   END_RUNG
   RUNG wire#w1
      Contact( %DB67.DBX7.1 )
      R_Coil( %DB60.DBX7.1 )
   END_RUNG
   RUNG wire#w1
      Contact( %DB67.DBX7.2 )
      R_Coil( %DB60.DBX7.2 )
   END_RUNG
   RUNG wire#w1
      Contact( %DB67.DBX7.3 )
      R_Coil( %DB60.DBX7.3 )
   END_RUNG
   RUNG wire#w1
      Contact( %DB67.DBX7.4 )
      R_Coil( %DB60.DBX7.4 )
   END_RUNG
   RUNG wire#w1
      Contact( %DB67.DBX7.5 )
      R_Coil( %DB60.DBX7.5 )
   END_RUNG
   RUNG wire#w1
      Contact( %DB67.DBX7.6 )
      R_Coil( %DB60.DBX7.6 )
   END_RUNG
   RUNG wire#w1
      Contact( %DB67.DBX7.7 )
      R_Coil( %DB60.DBX7.7 )
   END_RUNG
   // the same network as SCL:
   IF "AlwaysFALSE" AND %DB67.DBX0.0 THEN %DB60.DBX0.0 := FALSE; END_IF;
   IF "AlwaysFALSE" AND %DB67.DBX0.1 THEN %DB60.DBX0.1 := FALSE; END_IF;
   IF "AlwaysFALSE" AND %DB67.DBX0.2 THEN %DB60.DBX0.2 := FALSE; END_IF;
   IF "AlwaysFALSE" AND %DB67.DBX0.3 THEN %DB60.DBX0.3 := FALSE; END_IF;
   IF "AlwaysFALSE" AND %DB67.DBX0.4 THEN %DB60.DBX0.4 := FALSE; END_IF;
   IF "AlwaysFALSE" AND %DB67.DBX0.5 THEN %DB60.DBX0.5 := FALSE; END_IF;
   IF "AlwaysFALSE" AND %DB67.DBX0.6 THEN %DB60.DBX0.6 := FALSE; END_IF;
   IF "AlwaysFALSE" AND %DB67.DBX0.7 THEN %DB60.DBX0.7 := FALSE; END_IF;
   IF "AlwaysFALSE" AND %DB67.DBX1.0 THEN %DB60.DBX1.0 := FALSE; END_IF;
   IF "AlwaysFALSE" AND %DB67.DBX1.1 THEN %DB60.DBX1.1 := FALSE; END_IF;
   IF "AlwaysFALSE" AND %DB67.DBX1.2 THEN %DB60.DBX1.2 := FALSE; END_IF;
   IF "AlwaysFALSE" AND %DB67.DBX1.3 THEN %DB60.DBX1.3 := FALSE; END_IF;
   IF "AlwaysFALSE" AND %DB67.DBX1.4 THEN %DB60.DBX1.4 := FALSE; END_IF;
   IF "AlwaysFALSE" AND %DB67.DBX1.5 THEN %DB60.DBX1.5 := FALSE; END_IF;
   IF "AlwaysFALSE" AND %DB67.DBX1.6 THEN %DB60.DBX1.6 := FALSE; END_IF;
   IF "AlwaysFALSE" AND %DB67.DBX1.7 THEN %DB60.DBX1.7 := FALSE; END_IF;
   IF "AlwaysFALSE" AND %DB67.DBX2.0 THEN %DB60.DBX2.0 := FALSE; END_IF;
   IF "AlwaysFALSE" AND %DB67.DBX2.1 THEN %DB60.DBX2.1 := FALSE; END_IF;
   IF "AlwaysFALSE" AND %DB67.DBX2.2 THEN %DB60.DBX2.2 := FALSE; END_IF;
   IF "AlwaysFALSE" AND %DB67.DBX2.3 THEN %DB60.DBX2.3 := FALSE; END_IF;
   IF "AlwaysFALSE" AND %DB67.DBX2.4 THEN %DB60.DBX2.4 := FALSE; END_IF;
   IF "AlwaysFALSE" AND %DB67.DBX2.5 THEN %DB60.DBX2.5 := FALSE; END_IF;
   IF "AlwaysFALSE" AND %DB67.DBX2.6 THEN %DB60.DBX2.6 := FALSE; END_IF;
   IF "AlwaysFALSE" AND %DB67.DBX2.7 THEN %DB60.DBX2.7 := FALSE; END_IF;
   IF "AlwaysFALSE" AND %DB67.DBX3.0 THEN %DB60.DBX3.0 := FALSE; END_IF;
   IF "AlwaysFALSE" AND %DB67.DBX3.1 THEN %DB60.DBX3.1 := FALSE; END_IF;
   IF "AlwaysFALSE" AND %DB67.DBX3.2 THEN %DB60.DBX3.2 := FALSE; END_IF;
   IF "AlwaysFALSE" AND %DB67.DBX3.3 THEN %DB60.DBX3.3 := FALSE; END_IF;
   IF "AlwaysFALSE" AND %DB67.DBX3.4 THEN %DB60.DBX3.4 := FALSE; END_IF;
   IF "AlwaysFALSE" AND %DB67.DBX3.5 THEN %DB60.DBX3.5 := FALSE; END_IF;
   IF "AlwaysFALSE" AND %DB67.DBX3.6 THEN %DB60.DBX3.6 := FALSE; END_IF;
   IF "AlwaysFALSE" AND %DB67.DBX3.7 THEN %DB60.DBX3.7 := FALSE; END_IF;
   IF "AlwaysFALSE" AND %DB67.DBX4.0 THEN %DB60.DBX4.0 := FALSE; END_IF;
   IF "AlwaysFALSE" AND %DB67.DBX4.1 THEN %DB60.DBX4.1 := FALSE; END_IF;
   IF "AlwaysFALSE" AND %DB67.DBX4.2 THEN %DB60.DBX4.2 := FALSE; END_IF;
   IF "AlwaysFALSE" AND %DB67.DBX4.3 THEN %DB60.DBX4.3 := FALSE; END_IF;
   IF "AlwaysFALSE" AND %DB67.DBX4.4 THEN %DB60.DBX4.4 := FALSE; END_IF;
   IF "AlwaysFALSE" AND %DB67.DBX4.5 THEN %DB60.DBX4.5 := FALSE; END_IF;
   IF "AlwaysFALSE" AND %DB67.DBX4.6 THEN %DB60.DBX4.6 := FALSE; END_IF;
   IF "AlwaysFALSE" AND %DB67.DBX4.7 THEN %DB60.DBX4.7 := FALSE; END_IF;
   IF "AlwaysFALSE" AND %DB67.DBX5.0 THEN %DB60.DBX5.0 := FALSE; END_IF;
   IF "AlwaysFALSE" AND %DB67.DBX5.1 THEN %DB60.DBX5.1 := FALSE; END_IF;
   IF "AlwaysFALSE" AND %DB67.DBX5.2 THEN %DB60.DBX5.2 := FALSE; END_IF;
   IF "AlwaysFALSE" AND %DB67.DBX5.3 THEN %DB60.DBX5.3 := FALSE; END_IF;
   IF "AlwaysFALSE" AND %DB67.DBX5.4 THEN %DB60.DBX5.4 := FALSE; END_IF;
   IF "AlwaysFALSE" AND %DB67.DBX5.5 THEN %DB60.DBX5.5 := FALSE; END_IF;
   IF "AlwaysFALSE" AND %DB67.DBX5.6 THEN %DB60.DBX5.6 := FALSE; END_IF;
   IF "AlwaysFALSE" AND %DB67.DBX5.7 THEN %DB60.DBX5.7 := FALSE; END_IF;
   IF "AlwaysFALSE" AND %DB67.DBX6.0 THEN %DB60.DBX6.0 := FALSE; END_IF;
   IF "AlwaysFALSE" AND %DB67.DBX6.1 THEN %DB60.DBX6.1 := FALSE; END_IF;
   IF "AlwaysFALSE" AND %DB67.DBX6.2 THEN %DB60.DBX6.2 := FALSE; END_IF;
   IF "AlwaysFALSE" AND %DB67.DBX6.3 THEN %DB60.DBX6.3 := FALSE; END_IF;
   IF "AlwaysFALSE" AND %DB67.DBX6.4 THEN %DB60.DBX6.4 := FALSE; END_IF;
   IF "AlwaysFALSE" AND %DB67.DBX6.5 THEN %DB60.DBX6.5 := FALSE; END_IF;
   IF "AlwaysFALSE" AND %DB67.DBX6.6 THEN %DB60.DBX6.6 := FALSE; END_IF;
   IF "AlwaysFALSE" AND %DB67.DBX6.7 THEN %DB60.DBX6.7 := FALSE; END_IF;
   IF "AlwaysFALSE" AND %DB67.DBX7.0 THEN %DB60.DBX7.0 := FALSE; END_IF;
   IF "AlwaysFALSE" AND %DB67.DBX7.1 THEN %DB60.DBX7.1 := FALSE; END_IF;
   IF "AlwaysFALSE" AND %DB67.DBX7.2 THEN %DB60.DBX7.2 := FALSE; END_IF;
   IF "AlwaysFALSE" AND %DB67.DBX7.3 THEN %DB60.DBX7.3 := FALSE; END_IF;
   IF "AlwaysFALSE" AND %DB67.DBX7.4 THEN %DB60.DBX7.4 := FALSE; END_IF;
   IF "AlwaysFALSE" AND %DB67.DBX7.5 THEN %DB60.DBX7.5 := FALSE; END_IF;
   IF "AlwaysFALSE" AND %DB67.DBX7.6 THEN %DB60.DBX7.6 := FALSE; END_IF;
   IF "AlwaysFALSE" AND %DB67.DBX7.7 THEN %DB60.DBX7.7 := FALSE; END_IF;
END_REGION

REGION Network 48: Alarm Present
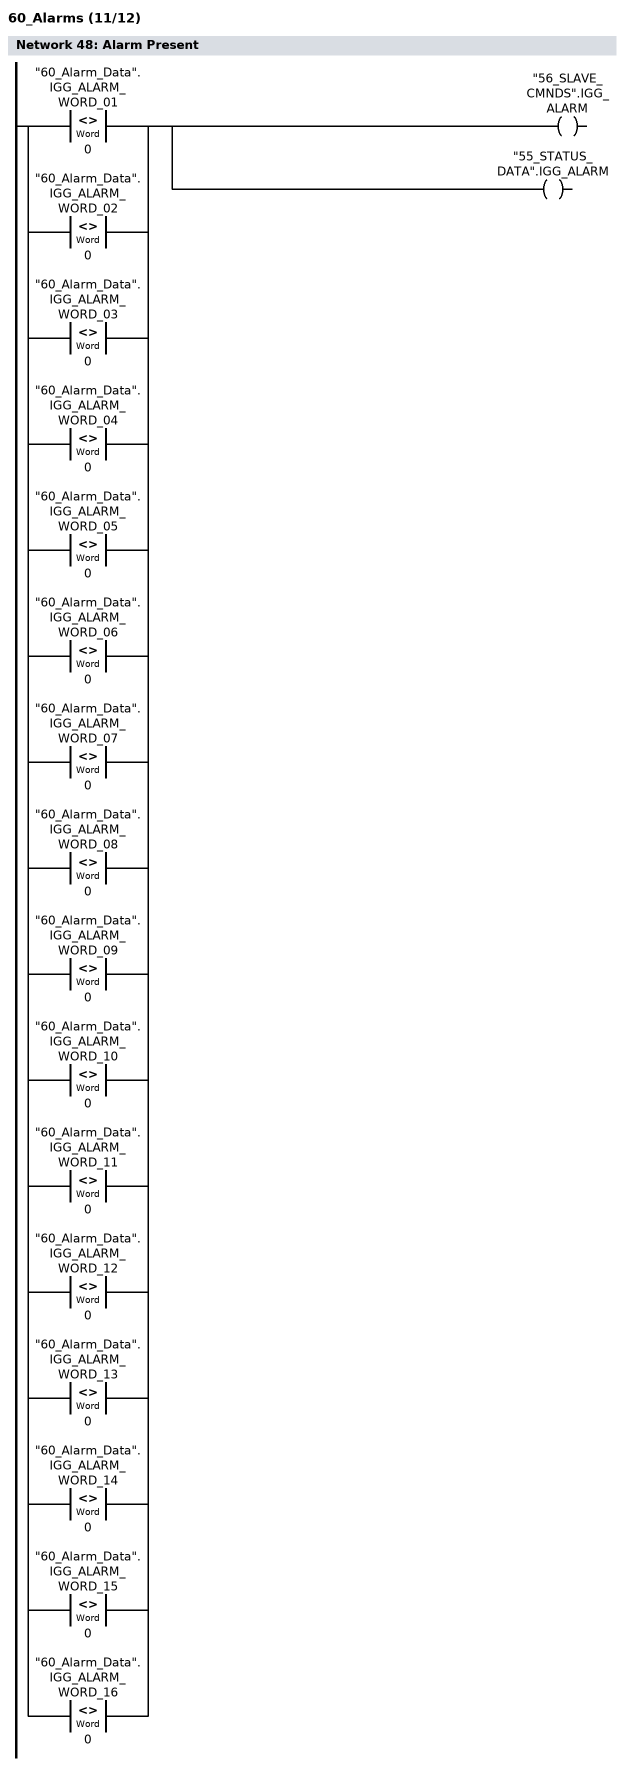
   RUNG wire#powerrail
      { S7_Templates := "SrcType := Word" } NE_Contact(in1 := "60_Alarm_Data".IGG_ALARM_WORD_01, in2 := 0)
      wire#w1
      Coil( "56_SLAVE_CMNDS".IGG_ALARM )
   END_RUNG
   RUNG wire#powerrail
      { S7_Templates := "SrcType := Word" } NE_Contact(in1 := "60_Alarm_Data".IGG_ALARM_WORD_02, in2 := 0)
   END_RUNG wire#w1
   RUNG wire#powerrail
      { S7_Templates := "SrcType := Word" } NE_Contact(in1 := "60_Alarm_Data".IGG_ALARM_WORD_03, in2 := 0)
   END_RUNG wire#w1
   RUNG wire#powerrail
      { S7_Templates := "SrcType := Word" } NE_Contact(in1 := "60_Alarm_Data".IGG_ALARM_WORD_04, in2 := 0)
   END_RUNG wire#w1
   RUNG wire#powerrail
      { S7_Templates := "SrcType := Word" } NE_Contact(in1 := "60_Alarm_Data".IGG_ALARM_WORD_05, in2 := 0)
   END_RUNG wire#w1
   RUNG wire#powerrail
      { S7_Templates := "SrcType := Word" } NE_Contact(in1 := "60_Alarm_Data".IGG_ALARM_WORD_06, in2 := 0)
   END_RUNG wire#w1
   RUNG wire#powerrail
      { S7_Templates := "SrcType := Word" } NE_Contact(in1 := "60_Alarm_Data".IGG_ALARM_WORD_07, in2 := 0)
   END_RUNG wire#w1
   RUNG wire#powerrail
      { S7_Templates := "SrcType := Word" } NE_Contact(in1 := "60_Alarm_Data".IGG_ALARM_WORD_08, in2 := 0)
   END_RUNG wire#w1
   RUNG wire#powerrail
      { S7_Templates := "SrcType := Word" } NE_Contact(in1 := "60_Alarm_Data".IGG_ALARM_WORD_09, in2 := 0)
   END_RUNG wire#w1
   RUNG wire#powerrail
      { S7_Templates := "SrcType := Word" } NE_Contact(in1 := "60_Alarm_Data".IGG_ALARM_WORD_10, in2 := 0)
   END_RUNG wire#w1
   RUNG wire#powerrail
      { S7_Templates := "SrcType := Word" } NE_Contact(in1 := "60_Alarm_Data".IGG_ALARM_WORD_11, in2 := 0)
   END_RUNG wire#w1
   RUNG wire#powerrail
      { S7_Templates := "SrcType := Word" } NE_Contact(in1 := "60_Alarm_Data".IGG_ALARM_WORD_12, in2 := 0)
   END_RUNG wire#w1
   RUNG wire#powerrail
      { S7_Templates := "SrcType := Word" } NE_Contact(in1 := "60_Alarm_Data".IGG_ALARM_WORD_13, in2 := 0)
   END_RUNG wire#w1
   RUNG wire#powerrail
      { S7_Templates := "SrcType := Word" } NE_Contact(in1 := "60_Alarm_Data".IGG_ALARM_WORD_14, in2 := 0)
   END_RUNG wire#w1
   RUNG wire#powerrail
      { S7_Templates := "SrcType := Word" } NE_Contact(in1 := "60_Alarm_Data".IGG_ALARM_WORD_15, in2 := 0)
   END_RUNG wire#w1
   RUNG wire#powerrail
      { S7_Templates := "SrcType := Word" } NE_Contact(in1 := "60_Alarm_Data".IGG_ALARM_WORD_16, in2 := 0)
   END_RUNG wire#w1
   RUNG wire#w1
      Coil( "55_STATUS_DATA".IGG_ALARM )
   END_RUNG
   // the same network as SCL:
   "56_SLAVE_CMNDS".IGG_ALARM := ("60_Alarm_Data".IGG_ALARM_WORD_01 <> 0) OR ("60_Alarm_Data".IGG_ALARM_WORD_02 <> 0) OR ("60_Alarm_Data".IGG_ALARM_WORD_03 <> 0) OR ("60_Alarm_Data".IGG_ALARM_WORD_04 <> 0) OR ("60_Alarm_Data".IGG_ALARM_WORD_05 <> 0) OR ("60_Alarm_Data".IGG_ALARM_WORD_06 <> 0) OR ("60_Alarm_Data".IGG_ALARM_WORD_07 <> 0) OR ("60_Alarm_Data".IGG_ALARM_WORD_08 <> 0) OR ("60_Alarm_Data".IGG_ALARM_WORD_09 <> 0) OR ("60_Alarm_Data".IGG_ALARM_WORD_10 <> 0) OR ("60_Alarm_Data".IGG_ALARM_WORD_11 <> 0) OR ("60_Alarm_Data".IGG_ALARM_WORD_12 <> 0) OR ("60_Alarm_Data".IGG_ALARM_WORD_13 <> 0) OR ("60_Alarm_Data".IGG_ALARM_WORD_14 <> 0) OR ("60_Alarm_Data".IGG_ALARM_WORD_15 <> 0) OR ("60_Alarm_Data".IGG_ALARM_WORD_16 <> 0);
   "55_STATUS_DATA".IGG_ALARM := "56_SLAVE_CMNDS".IGG_ALARM;
END_REGION

REGION Network 49: Alarm present
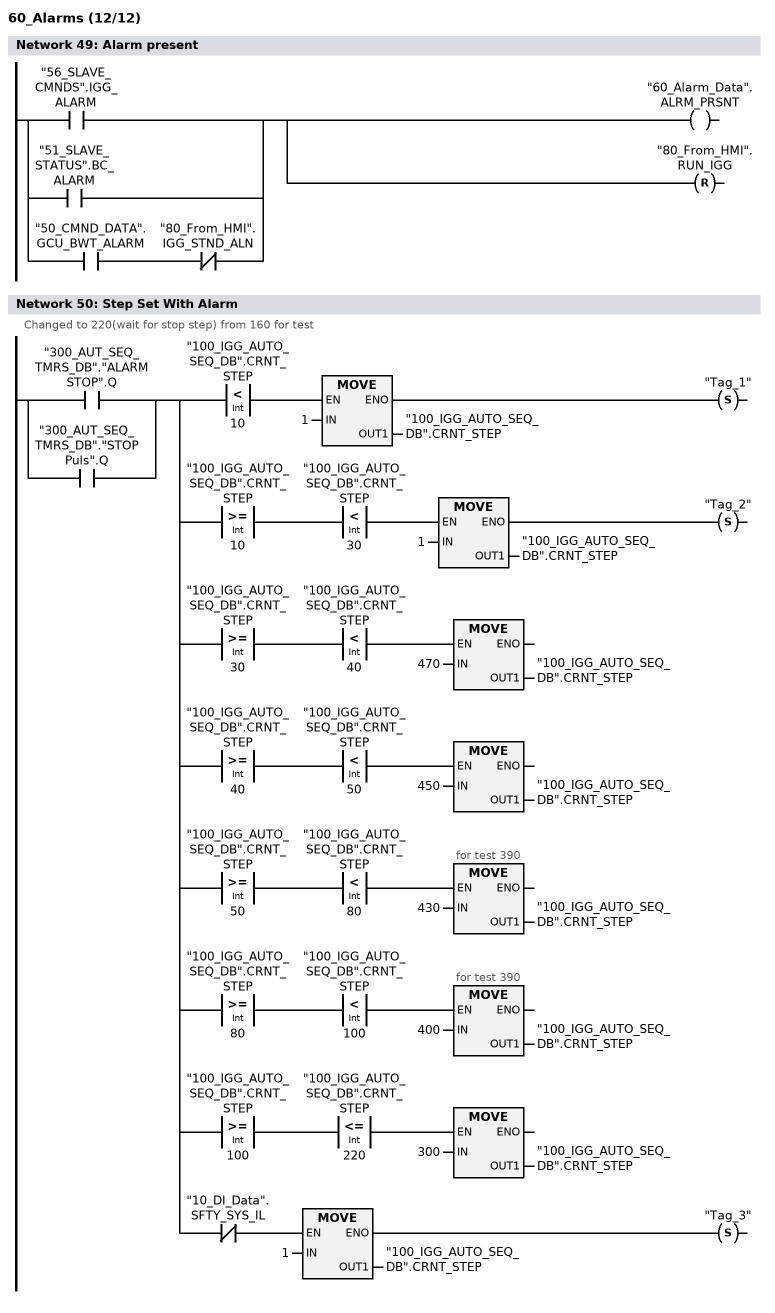
   RUNG wire#powerrail
      Contact( "56_SLAVE_CMNDS".IGG_ALARM )
      wire#w1
      Coil( "60_Alarm_Data".ALRM_PRSNT )
   END_RUNG
   RUNG wire#powerrail
      Contact( "51_SLAVE_STATUS".BC_ALARM )
   END_RUNG wire#w1
   RUNG wire#powerrail
      Contact( "50_CMND_DATA".GCU_BWT_ALARM )
      I_Contact( "80_From_HMI".IGG_STND_ALN )
   END_RUNG wire#w1
   RUNG wire#w1
      R_Coil( "80_From_HMI".RUN_IGG )
   END_RUNG
   // the same network as SCL:
   "60_Alarm_Data".ALRM_PRSNT := "56_SLAVE_CMNDS".IGG_ALARM OR "51_SLAVE_STATUS".BC_ALARM OR ("50_CMND_DATA".GCU_BWT_ALARM AND NOT "80_From_HMI".IGG_STND_ALN);
   IF "60_Alarm_Data".ALRM_PRSNT THEN "80_From_HMI".RUN_IGG := FALSE; END_IF;
END_REGION

REGION Network 50: Step Set With Alarm
   // Changed to 220(wait for stop step) from 160 for test
   RUNG wire#powerrail
      Contact( "300_AUT_SEQ_TMRS_DB"."ALARM STOP".Q )
      wire#w1
      { S7_Templates := "SrcType := Int" } LT_Contact(in1 := "100_IGG_AUTO_SEQ_DB".CRNT_STEP, in2 := 10)
      Move(in := 1, out1 => "100_IGG_AUTO_SEQ_DB".CRNT_STEP)
      S_Coil( "Tag_1" )
   END_RUNG
   RUNG wire#powerrail
      Contact( "300_AUT_SEQ_TMRS_DB"."STOP Puls".Q )
   END_RUNG wire#w1
   RUNG wire#w1
      { S7_Templates := "SrcType := Int" } GE_Contact(in1 := "100_IGG_AUTO_SEQ_DB".CRNT_STEP, in2 := 10)
      { S7_Templates := "SrcType := Int" } LT_Contact(in1 := "100_IGG_AUTO_SEQ_DB".CRNT_STEP, in2 := 30)
      Move(in := 1, out1 => "100_IGG_AUTO_SEQ_DB".CRNT_STEP)
      S_Coil( "Tag_2" )
   END_RUNG
   RUNG wire#w1
      { S7_Templates := "SrcType := Int" } GE_Contact(in1 := "100_IGG_AUTO_SEQ_DB".CRNT_STEP, in2 := 30)
      { S7_Templates := "SrcType := Int" } LT_Contact(in1 := "100_IGG_AUTO_SEQ_DB".CRNT_STEP, in2 := 40)
      Move(in := 470, out1 => "100_IGG_AUTO_SEQ_DB".CRNT_STEP)
   END_RUNG
   RUNG wire#w1
      { S7_Templates := "SrcType := Int" } GE_Contact(in1 := "100_IGG_AUTO_SEQ_DB".CRNT_STEP, in2 := 40)
      { S7_Templates := "SrcType := Int" } LT_Contact(in1 := "100_IGG_AUTO_SEQ_DB".CRNT_STEP, in2 := 50)
      Move(in := 450, out1 => "100_IGG_AUTO_SEQ_DB".CRNT_STEP)
   END_RUNG
   RUNG wire#w1
      { S7_Templates := "SrcType := Int" } GE_Contact(in1 := "100_IGG_AUTO_SEQ_DB".CRNT_STEP, in2 := 50)
      { S7_Templates := "SrcType := Int" } LT_Contact(in1 := "100_IGG_AUTO_SEQ_DB".CRNT_STEP, in2 := 80)
      Move(in := 430, out1 => "100_IGG_AUTO_SEQ_DB".CRNT_STEP)   // for test 390
   END_RUNG
   RUNG wire#w1
      { S7_Templates := "SrcType := Int" } GE_Contact(in1 := "100_IGG_AUTO_SEQ_DB".CRNT_STEP, in2 := 80)
      { S7_Templates := "SrcType := Int" } LT_Contact(in1 := "100_IGG_AUTO_SEQ_DB".CRNT_STEP, in2 := 100)
      Move(in := 400, out1 => "100_IGG_AUTO_SEQ_DB".CRNT_STEP)   // for test 390
   END_RUNG
   RUNG wire#w1
      { S7_Templates := "SrcType := Int" } GE_Contact(in1 := "100_IGG_AUTO_SEQ_DB".CRNT_STEP, in2 := 100)
      { S7_Templates := "SrcType := Int" } LE_Contact(in1 := "100_IGG_AUTO_SEQ_DB".CRNT_STEP, in2 := 220)
      Move(in := 300, out1 => "100_IGG_AUTO_SEQ_DB".CRNT_STEP)
   END_RUNG
   RUNG wire#w1
      I_Contact( "10_DI_Data".SFTY_SYS_IL )
      Move(in := 1, out1 => "100_IGG_AUTO_SEQ_DB".CRNT_STEP)
      S_Coil( "Tag_3" )
   END_RUNG
   // the same network as SCL:
   #_w1 := "300_AUT_SEQ_TMRS_DB"."ALARM STOP".Q OR "300_AUT_SEQ_TMRS_DB"."STOP Puls".Q;
   #_w2 := #_w1 AND ("100_IGG_AUTO_SEQ_DB".CRNT_STEP < 10);
   IF #_w2 THEN
       "100_IGG_AUTO_SEQ_DB".CRNT_STEP := 1;
       "Tag_1" := TRUE;
   END_IF;
   #_w3 := #_w1 AND ("100_IGG_AUTO_SEQ_DB".CRNT_STEP >= 10) AND ("100_IGG_AUTO_SEQ_DB".CRNT_STEP < 30);
   IF #_w3 THEN
       "100_IGG_AUTO_SEQ_DB".CRNT_STEP := 1;
       "Tag_2" := TRUE;
   END_IF;
   IF #_w1 AND ("100_IGG_AUTO_SEQ_DB".CRNT_STEP >= 30) AND ("100_IGG_AUTO_SEQ_DB".CRNT_STEP < 40) THEN
       "100_IGG_AUTO_SEQ_DB".CRNT_STEP := 470;
   END_IF;
   IF #_w1 AND ("100_IGG_AUTO_SEQ_DB".CRNT_STEP >= 40) AND ("100_IGG_AUTO_SEQ_DB".CRNT_STEP < 50) THEN
       "100_IGG_AUTO_SEQ_DB".CRNT_STEP := 450;
   END_IF;
   IF #_w1 AND ("100_IGG_AUTO_SEQ_DB".CRNT_STEP >= 50) AND ("100_IGG_AUTO_SEQ_DB".CRNT_STEP < 80) THEN
       "100_IGG_AUTO_SEQ_DB".CRNT_STEP := 430;   // for test 390
   END_IF;
   IF #_w1 AND ("100_IGG_AUTO_SEQ_DB".CRNT_STEP >= 80) AND ("100_IGG_AUTO_SEQ_DB".CRNT_STEP < 100) THEN
       "100_IGG_AUTO_SEQ_DB".CRNT_STEP := 400;   // for test 390
   END_IF;
   IF #_w1 AND ("100_IGG_AUTO_SEQ_DB".CRNT_STEP >= 100) AND ("100_IGG_AUTO_SEQ_DB".CRNT_STEP <= 220) THEN
       "100_IGG_AUTO_SEQ_DB".CRNT_STEP := 300;
   END_IF;
   IF #_w1 AND NOT "10_DI_Data".SFTY_SYS_IL THEN
       "100_IGG_AUTO_SEQ_DB".CRNT_STEP := 1;
       "Tag_3" := TRUE;
   END_IF;
END_REGION
END_FUNCTION

FUNCTION "62_Warnings" : Void   // FC62, LAD
TITLE = Warning Processing
{ S7_Optimized_Access := 'TRUE' }
AUTHOR : JRS
VERSION : 0.1
// To warning conditions
   VAR_TEMP   // added for the SCL form of the ladder/FBD networks
      _w1 : Bool;
   END_VAR
BEGIN

REGION Network 1: DB62 DBX0.0 = 31B1 Atmospheric O2 Sensor #1 O2
   // IGG_WARNING_WORD_01_BIT_0&2
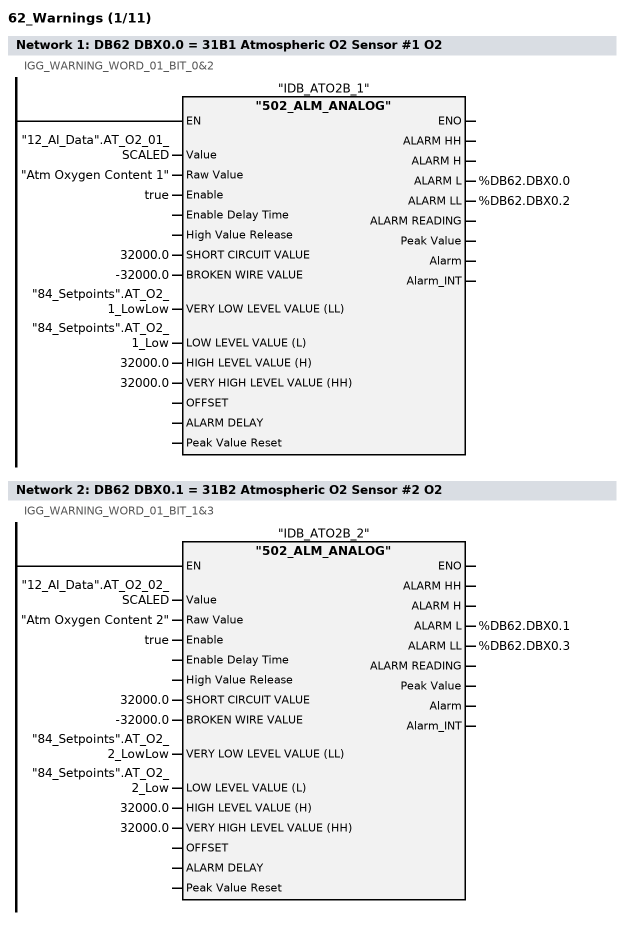
   RUNG wire#powerrail
      "IDB_ATO2B_1"(Value := "12_AI_Data".AT_O2_01_SCALED, "Raw Value" := "Atm Oxygen Content 1", Enable := true, "SHORT CIRCUIT VALUE" := 32000.0, "BROKEN WIRE VALUE" := -32000.0, "VERY LOW LEVEL VALUE (LL)" := "84_Setpoints".AT_O2_1_LowLow, "LOW LEVEL VALUE (L)" := "84_Setpoints".AT_O2_1_Low, "HIGH LEVEL VALUE (H)" := 32000.0, "VERY HIGH LEVEL VALUE (HH)" := 32000.0, OFFSET :=, "ALARM DELAY" :=, "Peak Value Reset" :=, "ALARM HH" =>, "ALARM H" =>, "ALARM L" => %DB62.DBX0.0, "ALARM LL" => %DB62.DBX0.2, "ALARM READING" =>, "Peak Value" =>, Alarm =>, Alarm_INT =>, "Enable Delay Time" :=, "High Value Release" :=)
   END_RUNG
   // the same network as SCL:
   "IDB_ATO2B_1"(Value := "12_AI_Data".AT_O2_01_SCALED,   // "502_ALM_ANALOG"
                 "Raw Value" := "Atm Oxygen Content 1",
                 Enable := true,
                 "SHORT CIRCUIT VALUE" := 32000.0,
                 "BROKEN WIRE VALUE" := -32000.0,
                 "VERY LOW LEVEL VALUE (LL)" := "84_Setpoints".AT_O2_1_LowLow,
                 "LOW LEVEL VALUE (L)" := "84_Setpoints".AT_O2_1_Low,
                 "HIGH LEVEL VALUE (H)" := 32000.0,
                 "VERY HIGH LEVEL VALUE (HH)" := 32000.0,
                 "ALARM L" => %DB62.DBX0.0,
                 "ALARM LL" => %DB62.DBX0.2);
END_REGION

REGION Network 2: DB62 DBX0.1 = 31B2 Atmospheric O2 Sensor #2 O2
   // IGG_WARNING_WORD_01_BIT_1&3
   RUNG wire#powerrail
      "IDB_ATO2B_2"(Value := "12_AI_Data".AT_O2_02_SCALED, "Raw Value" := "Atm Oxygen Content 2", Enable := true, "SHORT CIRCUIT VALUE" := 32000.0, "BROKEN WIRE VALUE" := -32000.0, "VERY LOW LEVEL VALUE (LL)" := "84_Setpoints".AT_O2_2_LowLow, "LOW LEVEL VALUE (L)" := "84_Setpoints".AT_O2_2_Low, "HIGH LEVEL VALUE (H)" := 32000.0, "VERY HIGH LEVEL VALUE (HH)" := 32000.0, OFFSET :=, "ALARM DELAY" :=, "Peak Value Reset" :=, "ALARM HH" =>, "ALARM H" =>, "ALARM L" => %DB62.DBX0.1, "ALARM LL" => %DB62.DBX0.3, "ALARM READING" =>, "Peak Value" =>, Alarm =>, Alarm_INT =>, "Enable Delay Time" :=, "High Value Release" :=)
   END_RUNG
   // the same network as SCL:
   "IDB_ATO2B_2"(Value := "12_AI_Data".AT_O2_02_SCALED,   // "502_ALM_ANALOG"
                 "Raw Value" := "Atm Oxygen Content 2",
                 Enable := true,
                 "SHORT CIRCUIT VALUE" := 32000.0,
                 "BROKEN WIRE VALUE" := -32000.0,
                 "VERY LOW LEVEL VALUE (LL)" := "84_Setpoints".AT_O2_2_LowLow,
                 "LOW LEVEL VALUE (L)" := "84_Setpoints".AT_O2_2_Low,
                 "HIGH LEVEL VALUE (H)" := 32000.0,
                 "VERY HIGH LEVEL VALUE (HH)" := 32000.0,
                 "ALARM L" => %DB62.DBX0.1,
                 "ALARM LL" => %DB62.DBX0.3);
END_REGION

REGION Network 4: DB62 DBX2.0/2.1/5.0/5.1 = PIT102 CA Pressure
   // IGG_WARNING_WORD_02&03_BIT_0&1
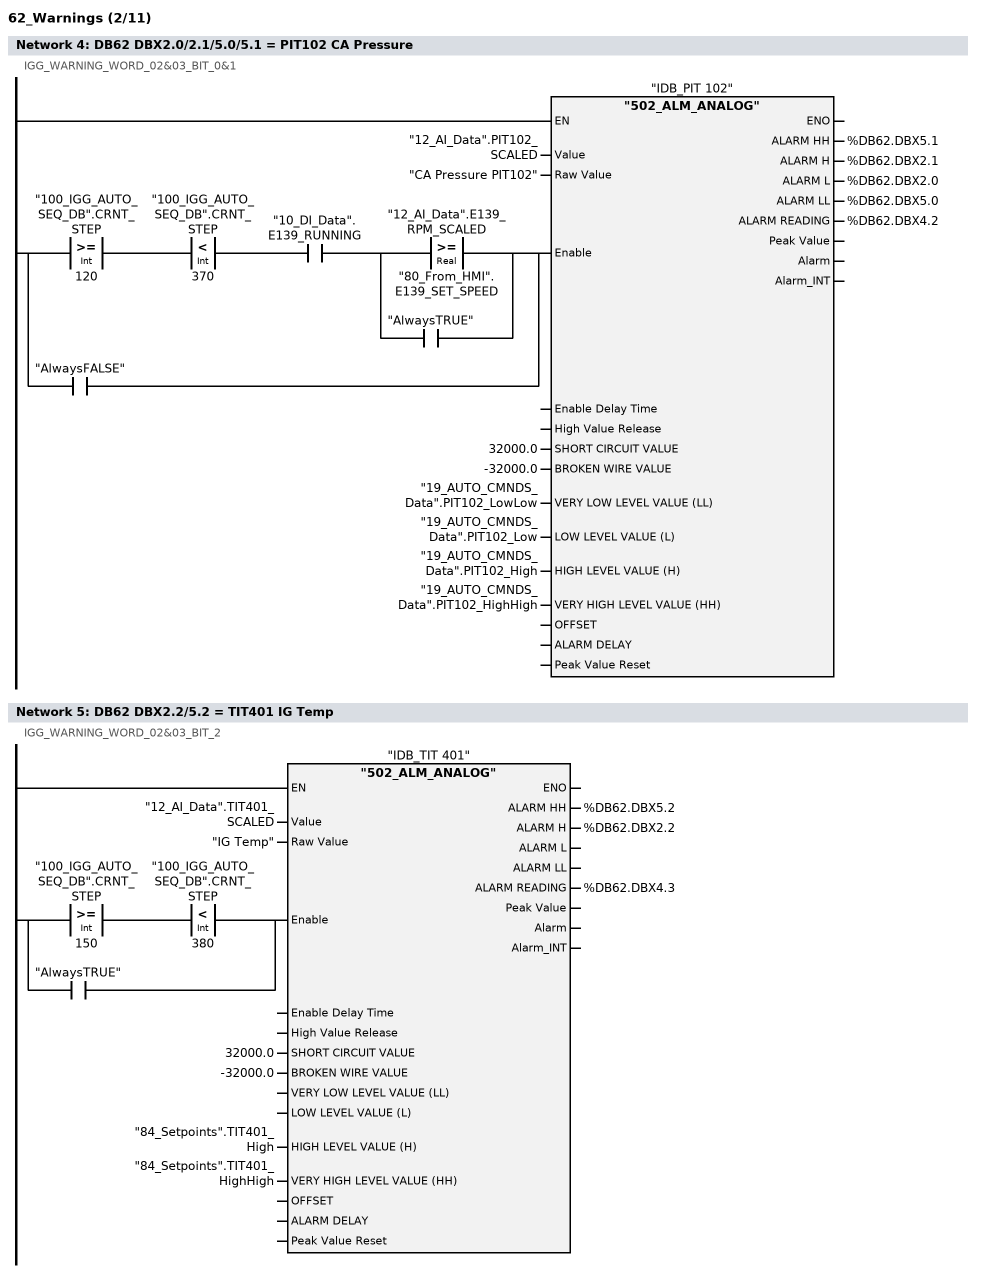
   RUNG wire#powerrail
      "IDB_PIT 102"(Enable := wire#w2, Value := "12_AI_Data".PIT102_SCALED, "Raw Value" := "CA Pressure PIT102", "SHORT CIRCUIT VALUE" := 32000.0, "BROKEN WIRE VALUE" := -32000.0, "VERY LOW LEVEL VALUE (LL)" := "19_AUTO_CMNDS_Data".PIT102_LowLow, "LOW LEVEL VALUE (L)" := "19_AUTO_CMNDS_Data".PIT102_Low, "HIGH LEVEL VALUE (H)" := "19_AUTO_CMNDS_Data".PIT102_High, "VERY HIGH LEVEL VALUE (HH)" := "19_AUTO_CMNDS_Data".PIT102_HighHigh, OFFSET :=, "ALARM DELAY" :=, "Peak Value Reset" :=, "ALARM HH" => %DB62.DBX5.1, "ALARM H" => %DB62.DBX2.1, "ALARM L" => %DB62.DBX2.0, "ALARM LL" => %DB62.DBX5.0, "ALARM READING" => %DB62.DBX4.2, "Peak Value" =>, Alarm =>, Alarm_INT =>, "Enable Delay Time" :=, "High Value Release" :=)
   END_RUNG
   RUNG wire#powerrail
      { S7_Templates := "SrcType := Int" } GE_Contact(in1 := "100_IGG_AUTO_SEQ_DB".CRNT_STEP, in2 := 120)
      { S7_Templates := "SrcType := Int" } LT_Contact(in1 := "100_IGG_AUTO_SEQ_DB".CRNT_STEP, in2 := 370)
      Contact( "10_DI_Data".E139_RUNNING )
      wire#w1
      { S7_Templates := "SrcType := Real" } GE_Contact(in1 := "12_AI_Data".E139_RPM_SCALED, in2 := "80_From_HMI".E139_SET_SPEED)
   END_RUNG wire#w2
   RUNG wire#w1
      Contact( "AlwaysTRUE" )
   END_RUNG wire#w2
   RUNG wire#powerrail
      Contact( "AlwaysFALSE" )
   END_RUNG wire#w2
   // the same network as SCL:
   "IDB_PIT 102"(Value := "12_AI_Data".PIT102_SCALED,   // "502_ALM_ANALOG"
                 "Raw Value" := "CA Pressure PIT102",
                 Enable := (("100_IGG_AUTO_SEQ_DB".CRNT_STEP >= 120) AND ("100_IGG_AUTO_SEQ_DB".CRNT_STEP < 370) AND "10_DI_Data".E139_RUNNING AND (("12_AI_Data".E139_RPM_SCALED >= "80_From_HMI".E139_SET_SPEED) OR "AlwaysTRUE")) OR "AlwaysFALSE",
                 "SHORT CIRCUIT VALUE" := 32000.0,
                 "BROKEN WIRE VALUE" := -32000.0,
                 "VERY LOW LEVEL VALUE (LL)" := "19_AUTO_CMNDS_Data".PIT102_LowLow,
                 "LOW LEVEL VALUE (L)" := "19_AUTO_CMNDS_Data".PIT102_Low,
                 "HIGH LEVEL VALUE (H)" := "19_AUTO_CMNDS_Data".PIT102_High,
                 "VERY HIGH LEVEL VALUE (HH)" := "19_AUTO_CMNDS_Data".PIT102_HighHigh,
                 "ALARM HH" => %DB62.DBX5.1,
                 "ALARM H" => %DB62.DBX2.1,
                 "ALARM L" => %DB62.DBX2.0,
                 "ALARM LL" => %DB62.DBX5.0,
                 "ALARM READING" => %DB62.DBX4.2);
END_REGION

REGION Network 5: DB62 DBX2.2/5.2 = TIT401 IG Temp
   // IGG_WARNING_WORD_02&03_BIT_2
   RUNG wire#powerrail
      "IDB_TIT 401"(Enable := wire#w1, Value := "12_AI_Data".TIT401_SCALED, "Raw Value" := "IG Temp", "SHORT CIRCUIT VALUE" := 32000.0, "BROKEN WIRE VALUE" := -32000.0, "VERY LOW LEVEL VALUE (LL)" :=, "LOW LEVEL VALUE (L)" :=, "HIGH LEVEL VALUE (H)" := "84_Setpoints".TIT401_High, "VERY HIGH LEVEL VALUE (HH)" := "84_Setpoints".TIT401_HighHigh, OFFSET :=, "ALARM DELAY" :=, "Peak Value Reset" :=, "ALARM HH" => %DB62.DBX5.2, "ALARM H" => %DB62.DBX2.2, "ALARM L" =>, "ALARM LL" =>, "ALARM READING" => %DB62.DBX4.3, "Peak Value" =>, Alarm =>, Alarm_INT =>, "Enable Delay Time" :=, "High Value Release" :=)
   END_RUNG
   RUNG wire#powerrail
      { S7_Templates := "SrcType := Int" } GE_Contact(in1 := "100_IGG_AUTO_SEQ_DB".CRNT_STEP, in2 := 150)
      { S7_Templates := "SrcType := Int" } LT_Contact(in1 := "100_IGG_AUTO_SEQ_DB".CRNT_STEP, in2 := 380)
   END_RUNG wire#w1
   RUNG wire#powerrail
      Contact( "AlwaysTRUE" )
   END_RUNG wire#w1
   // the same network as SCL:
   "IDB_TIT 401"(Value := "12_AI_Data".TIT401_SCALED,   // "502_ALM_ANALOG"
                 "Raw Value" := "IG Temp",
                 Enable := (("100_IGG_AUTO_SEQ_DB".CRNT_STEP >= 150) AND ("100_IGG_AUTO_SEQ_DB".CRNT_STEP < 380)) OR "AlwaysTRUE",
                 "SHORT CIRCUIT VALUE" := 32000.0,
                 "BROKEN WIRE VALUE" := -32000.0,
                 "HIGH LEVEL VALUE (H)" := "84_Setpoints".TIT401_High,
                 "VERY HIGH LEVEL VALUE (HH)" := "84_Setpoints".TIT401_HighHigh,
                 "ALARM HH" => %DB62.DBX5.2,
                 "ALARM H" => %DB62.DBX2.2,
                 "ALARM READING" => %DB62.DBX4.3);
END_REGION

REGION Network 6: DB62 DBX2.3/2.4/5.3/5.4 = PIT402
   // IGG_WARNING_WORD_02&03_BIT_3&4
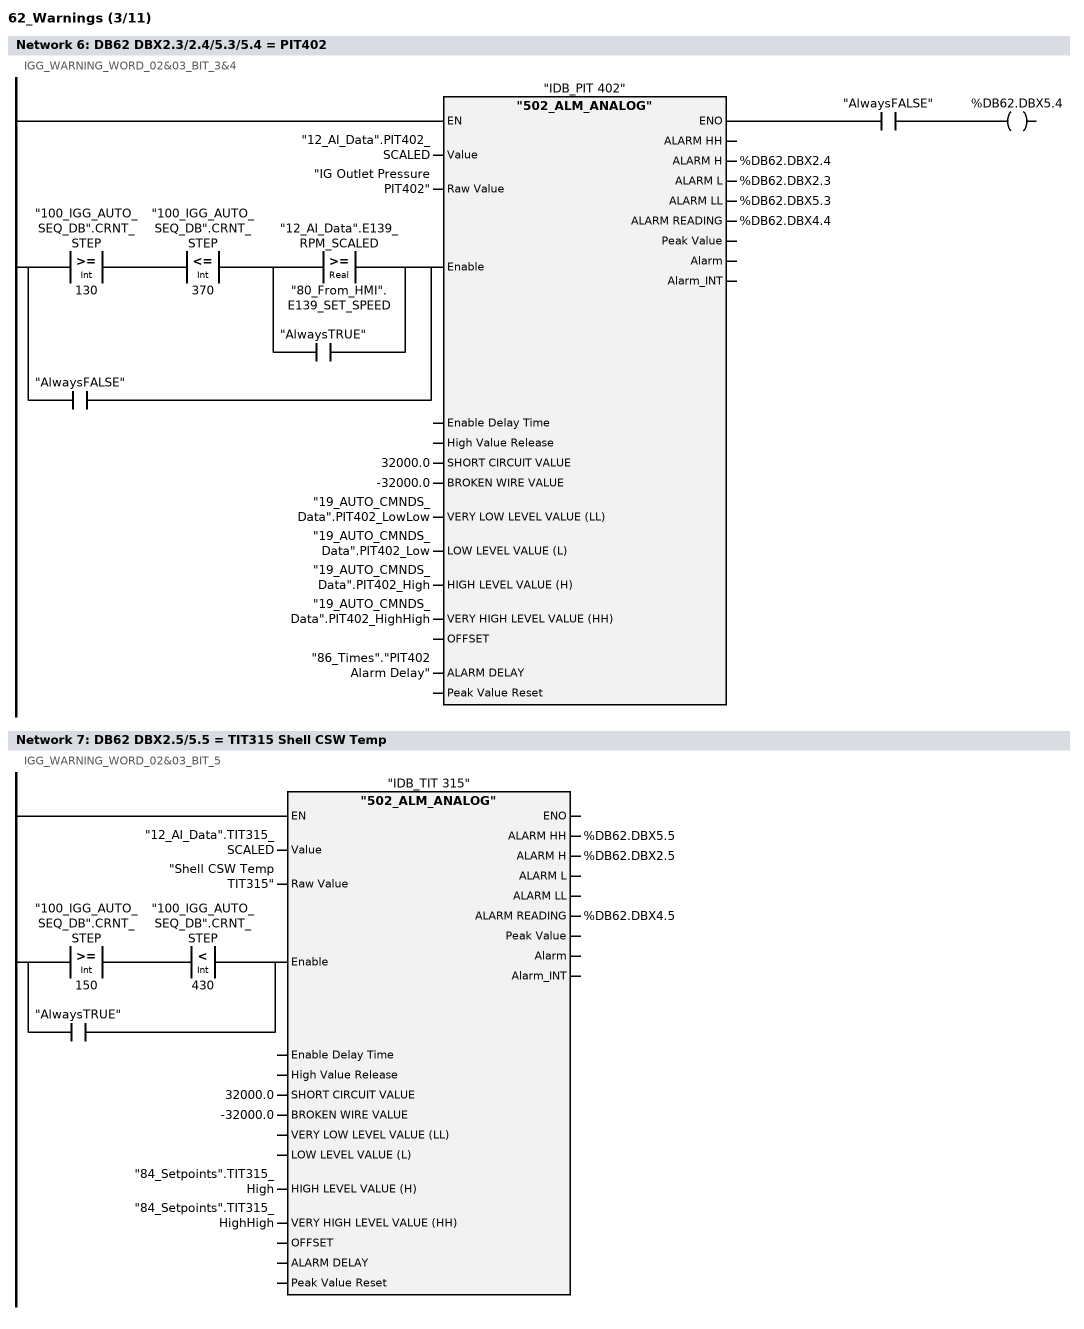
   RUNG wire#powerrail
      "IDB_PIT 402"(Enable := wire#w2, Value := "12_AI_Data".PIT402_SCALED, "Raw Value" := "IG Outlet Pressure PIT402", "Enable Delay Time" :=, "High Value Release" :=, "SHORT CIRCUIT VALUE" := 32000.0, "BROKEN WIRE VALUE" := -32000.0, "VERY LOW LEVEL VALUE (LL)" := "19_AUTO_CMNDS_Data".PIT402_LowLow, "LOW LEVEL VALUE (L)" := "19_AUTO_CMNDS_Data".PIT402_Low, "HIGH LEVEL VALUE (H)" := "19_AUTO_CMNDS_Data".PIT402_High, "VERY HIGH LEVEL VALUE (HH)" := "19_AUTO_CMNDS_Data".PIT402_HighHigh, OFFSET :=, "ALARM DELAY" := "86_Times"."PIT402 Alarm Delay", "Peak Value Reset" :=, "ALARM HH" =>, "ALARM H" => %DB62.DBX2.4, "ALARM L" => %DB62.DBX2.3, "ALARM LL" => %DB62.DBX5.3, "ALARM READING" => %DB62.DBX4.4, "Peak Value" =>, Alarm =>, Alarm_INT =>)
      Contact( "AlwaysFALSE" )
      Coil( %DB62.DBX5.4 )
   END_RUNG
   RUNG wire#powerrail
      { S7_Templates := "SrcType := Int" } GE_Contact(in1 := "100_IGG_AUTO_SEQ_DB".CRNT_STEP, in2 := 130)
      { S7_Templates := "SrcType := Int" } LE_Contact(in1 := "100_IGG_AUTO_SEQ_DB".CRNT_STEP, in2 := 370)
      wire#w1
      { S7_Templates := "SrcType := Real" } GE_Contact(in1 := "12_AI_Data".E139_RPM_SCALED, in2 := "80_From_HMI".E139_SET_SPEED)
   END_RUNG wire#w2
   RUNG wire#w1
      Contact( "AlwaysTRUE" )
   END_RUNG wire#w2
   RUNG wire#powerrail
      Contact( "AlwaysFALSE" )
   END_RUNG wire#w2
   // the same network as SCL:
   "IDB_PIT 402"(Value := "12_AI_Data".PIT402_SCALED,   // "502_ALM_ANALOG"
                 "Raw Value" := "IG Outlet Pressure PIT402",
                 Enable := (("100_IGG_AUTO_SEQ_DB".CRNT_STEP >= 130) AND ("100_IGG_AUTO_SEQ_DB".CRNT_STEP <= 370) AND (("12_AI_Data".E139_RPM_SCALED >= "80_From_HMI".E139_SET_SPEED) OR "AlwaysTRUE")) OR "AlwaysFALSE",
                 "SHORT CIRCUIT VALUE" := 32000.0,
                 "BROKEN WIRE VALUE" := -32000.0,
                 "VERY LOW LEVEL VALUE (LL)" := "19_AUTO_CMNDS_Data".PIT402_LowLow,
                 "LOW LEVEL VALUE (L)" := "19_AUTO_CMNDS_Data".PIT402_Low,
                 "HIGH LEVEL VALUE (H)" := "19_AUTO_CMNDS_Data".PIT402_High,
                 "VERY HIGH LEVEL VALUE (HH)" := "19_AUTO_CMNDS_Data".PIT402_HighHigh,
                 "ALARM DELAY" := "86_Times"."PIT402 Alarm Delay",
                 "ALARM H" => %DB62.DBX2.4,
                 "ALARM L" => %DB62.DBX2.3,
                 "ALARM LL" => %DB62.DBX5.3,
                 "ALARM READING" => %DB62.DBX4.4,
                 ENO => #_w1);
   %DB62.DBX5.4 := #_w1 AND "AlwaysFALSE";
END_REGION

REGION Network 7: DB62 DBX2.5/5.5 = TIT315 Shell CSW Temp
   // IGG_WARNING_WORD_02&03_BIT_5
   RUNG wire#powerrail
      "IDB_TIT 315"(Enable := wire#w1, Value := "12_AI_Data".TIT315_SCALED, "Raw Value" := "Shell CSW Temp TIT315", "SHORT CIRCUIT VALUE" := 32000.0, "BROKEN WIRE VALUE" := -32000.0, "VERY LOW LEVEL VALUE (LL)" :=, "LOW LEVEL VALUE (L)" :=, "HIGH LEVEL VALUE (H)" := "84_Setpoints".TIT315_High, "VERY HIGH LEVEL VALUE (HH)" := "84_Setpoints".TIT315_HighHigh, OFFSET :=, "ALARM DELAY" :=, "Peak Value Reset" :=, "ALARM HH" => %DB62.DBX5.5, "ALARM H" => %DB62.DBX2.5, "ALARM L" =>, "ALARM LL" =>, "ALARM READING" => %DB62.DBX4.5, "Peak Value" =>, Alarm =>, Alarm_INT =>, "Enable Delay Time" :=, "High Value Release" :=)
   END_RUNG
   RUNG wire#powerrail
      { S7_Templates := "SrcType := Int" } GE_Contact(in1 := "100_IGG_AUTO_SEQ_DB".CRNT_STEP, in2 := 150)
      { S7_Templates := "SrcType := Int" } LT_Contact(in1 := "100_IGG_AUTO_SEQ_DB".CRNT_STEP, in2 := 430)
   END_RUNG wire#w1
   RUNG wire#powerrail
      Contact( "AlwaysTRUE" )
   END_RUNG wire#w1
   // the same network as SCL:
   "IDB_TIT 315"(Value := "12_AI_Data".TIT315_SCALED,   // "502_ALM_ANALOG"
                 "Raw Value" := "Shell CSW Temp TIT315",
                 Enable := (("100_IGG_AUTO_SEQ_DB".CRNT_STEP >= 150) AND ("100_IGG_AUTO_SEQ_DB".CRNT_STEP < 430)) OR "AlwaysTRUE",
                 "SHORT CIRCUIT VALUE" := 32000.0,
                 "BROKEN WIRE VALUE" := -32000.0,
                 "HIGH LEVEL VALUE (H)" := "84_Setpoints".TIT315_High,
                 "VERY HIGH LEVEL VALUE (HH)" := "84_Setpoints".TIT315_HighHigh,
                 "ALARM HH" => %DB62.DBX5.5,
                 "ALARM H" => %DB62.DBX2.5,
                 "ALARM READING" => %DB62.DBX4.5);
END_REGION

REGION Network 8: DB62 DBX2.6/5.6 = TIT319 Inlet CSW Temp
   // IGG_WARNING_WORD_02&03_BIT_6